REGION Network 7
   // *********************************************************************************************************************
   // 
   // Next Carrier Traffic Cop Motion Function Block FB111. Traffic Cop and carrier motion logic for Zone called in Function block call located  in OB1.  Function block contains logic for Motion control and Traffic Cop logic for Carrier located in Position 3 of called Zone.  Carrier position within the zone is contained in the Tag    - “ Zone.[called zone].CarrierZnStatus[Position in zone].  Input parameter “MaxCarriers” Zones are divided into positions based on “MaxCarriers” allowed in zone which is set in the zone setup function block and represents the maximum number of carriers within the zone. 
   // 
   // **********************************************************************************************************************
   RUNG wire#powerrail
      "IDB602_NextCarrierTCopMotionFB"(Zone := #Zone, ZonePos := 3, CarrierNumber => "DB116_TC_ZoneMotionControl".Zone[#Zone].ZonePos[3].CarrierNumber, MoveFwdCommand => "DB116_TC_ZoneMotionControl".Zone[#Zone].ZonePos[3].MoveFwd, DriveCmdSpeed => "DB116_TC_ZoneMotionControl".Zone[#Zone].ZonePos[3].DriveCmdSpeed, NextStopPosition => "DB116_TC_ZoneMotionControl".Zone[#Zone].ZonePos[3].NextStopPos, NextCarrierNum => "DB116_TC_ZoneMotionControl".Zone[#Zone].ZonePos[3].NextCarrierNumber, AtCmdPosition => "DB116_TC_ZoneMotionControl".Zone[#Zone].ZonePos[3].AtCmdPos)
   END_RUNG
   // the same network as SCL:
   "IDB602_NextCarrierTCopMotionFB"(Zone := #Zone,   // "FB111_NextCarrierTCopMotionFB"
                           ZonePos := 3,
                           CarrierNumber => "DB116_TC_ZoneMotionControl".Zone[#Zone].ZonePos[3].CarrierNumber,
                           MoveFwdCommand => "DB116_TC_ZoneMotionControl".Zone[#Zone].ZonePos[3].MoveFwd,
                           DriveCmdSpeed => "DB116_TC_ZoneMotionControl".Zone[#Zone].ZonePos[3].DriveCmdSpeed,
                           NextStopPosition => "DB116_TC_ZoneMotionControl".Zone[#Zone].ZonePos[3].NextStopPos,
                           NextCarrierNum => "DB116_TC_ZoneMotionControl".Zone[#Zone].ZonePos[3].NextCarrierNumber,
                           AtCmdPosition => "DB116_TC_ZoneMotionControl".Zone[#Zone].ZonePos[3].AtCmdPos);
END_REGION

REGION Network 8
   // *********************************************************************************************************************
   // 
   // Next Carrier Traffic Cop Motion Function Block FB111. Traffic Cop and carrier motion logic for Zone called in Function block call located  in OB1.  Function block contains logic for Motion control and Traffic Cop logic for Carrier located in Position 4 of called Zone.  Carrier position within the zone is contained in the Tag    - “ Zone.[called zone].CarrierZnStatus[Position in zone].  Input parameter “MaxCarriers” Zones are divided into positions based on “MaxCarriers” allowed in zone which is set in the zone setup function block and represents the maximum number of carriers within the zone. 
   // 
   // **********************************************************************************************************************
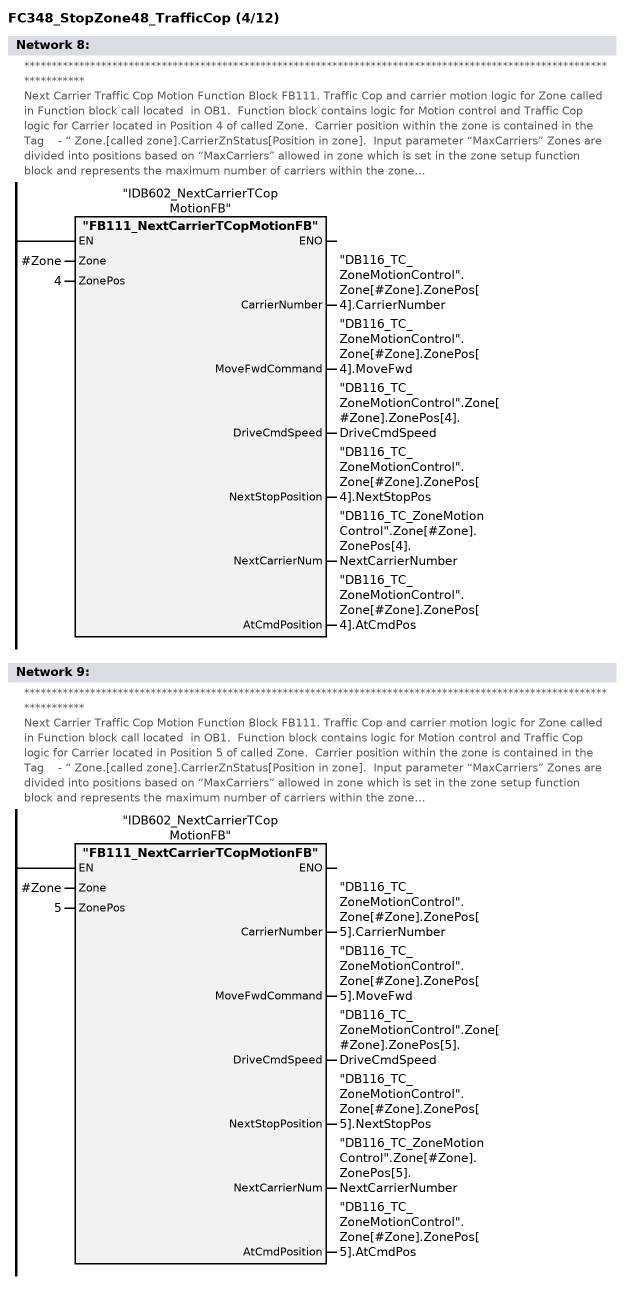
   RUNG wire#powerrail
      "IDB602_NextCarrierTCopMotionFB"(Zone := #Zone, ZonePos := 4, CarrierNumber => "DB116_TC_ZoneMotionControl".Zone[#Zone].ZonePos[4].CarrierNumber, MoveFwdCommand => "DB116_TC_ZoneMotionControl".Zone[#Zone].ZonePos[4].MoveFwd, DriveCmdSpeed => "DB116_TC_ZoneMotionControl".Zone[#Zone].ZonePos[4].DriveCmdSpeed, NextStopPosition => "DB116_TC_ZoneMotionControl".Zone[#Zone].ZonePos[4].NextStopPos, NextCarrierNum => "DB116_TC_ZoneMotionControl".Zone[#Zone].ZonePos[4].NextCarrierNumber, AtCmdPosition => "DB116_TC_ZoneMotionControl".Zone[#Zone].ZonePos[4].AtCmdPos)
   END_RUNG
   // the same network as SCL:
   "IDB602_NextCarrierTCopMotionFB"(Zone := #Zone,   // "FB111_NextCarrierTCopMotionFB"
                           ZonePos := 4,
                           CarrierNumber => "DB116_TC_ZoneMotionControl".Zone[#Zone].ZonePos[4].CarrierNumber,
                           MoveFwdCommand => "DB116_TC_ZoneMotionControl".Zone[#Zone].ZonePos[4].MoveFwd,
                           DriveCmdSpeed => "DB116_TC_ZoneMotionControl".Zone[#Zone].ZonePos[4].DriveCmdSpeed,
                           NextStopPosition => "DB116_TC_ZoneMotionControl".Zone[#Zone].ZonePos[4].NextStopPos,
                           NextCarrierNum => "DB116_TC_ZoneMotionControl".Zone[#Zone].ZonePos[4].NextCarrierNumber,
                           AtCmdPosition => "DB116_TC_ZoneMotionControl".Zone[#Zone].ZonePos[4].AtCmdPos);
END_REGION

REGION Network 9
   // *********************************************************************************************************************
   // 
   // Next Carrier Traffic Cop Motion Function Block FB111. Traffic Cop and carrier motion logic for Zone called in Function block call located  in OB1.  Function block contains logic for Motion control and Traffic Cop logic for Carrier located in Position 5 of called Zone.  Carrier position within the zone is contained in the Tag    - “ Zone.[called zone].CarrierZnStatus[Position in zone].  Input parameter “MaxCarriers” Zones are divided into positions based on “MaxCarriers” allowed in zone which is set in the zone setup function block and represents the maximum number of carriers within the zone. 
   // 
   // **********************************************************************************************************************
   RUNG wire#powerrail
      "IDB602_NextCarrierTCopMotionFB"(Zone := #Zone, ZonePos := 5, CarrierNumber => "DB116_TC_ZoneMotionControl".Zone[#Zone].ZonePos[5].CarrierNumber, MoveFwdCommand => "DB116_TC_ZoneMotionControl".Zone[#Zone].ZonePos[5].MoveFwd, DriveCmdSpeed => "DB116_TC_ZoneMotionControl".Zone[#Zone].ZonePos[5].DriveCmdSpeed, NextStopPosition => "DB116_TC_ZoneMotionControl".Zone[#Zone].ZonePos[5].NextStopPos, NextCarrierNum => "DB116_TC_ZoneMotionControl".Zone[#Zone].ZonePos[5].NextCarrierNumber, AtCmdPosition => "DB116_TC_ZoneMotionControl".Zone[#Zone].ZonePos[5].AtCmdPos)
   END_RUNG
   // the same network as SCL:
   "IDB602_NextCarrierTCopMotionFB"(Zone := #Zone,   // "FB111_NextCarrierTCopMotionFB"
                           ZonePos := 5,
                           CarrierNumber => "DB116_TC_ZoneMotionControl".Zone[#Zone].ZonePos[5].CarrierNumber,
                           MoveFwdCommand => "DB116_TC_ZoneMotionControl".Zone[#Zone].ZonePos[5].MoveFwd,
                           DriveCmdSpeed => "DB116_TC_ZoneMotionControl".Zone[#Zone].ZonePos[5].DriveCmdSpeed,
                           NextStopPosition => "DB116_TC_ZoneMotionControl".Zone[#Zone].ZonePos[5].NextStopPos,
                           NextCarrierNum => "DB116_TC_ZoneMotionControl".Zone[#Zone].ZonePos[5].NextCarrierNumber,
                           AtCmdPosition => "DB116_TC_ZoneMotionControl".Zone[#Zone].ZonePos[5].AtCmdPos);
END_REGION

REGION Network 10
   // *********************************************************************************************************************
   // 
   // Next Carrier Traffic Cop Motion Function Block FB111. Traffic Cop and carrier motion logic for Zone called in Function block call located  in OB1.  Function block contains logic for Motion control and Traffic Cop logic for Carrier located in Position 6 of called Zone.  Carrier position within the zone is contained in the Tag    - “ Zone.[called zone].CarrierZnStatus[Position in zone].  Input parameter “MaxCarriers” Zones are divided into positions based on “MaxCarriers” allowed in zone which is set in the zone setup function block and represents the maximum number of carriers within the zone. 
   // 
   // **********************************************************************************************************************
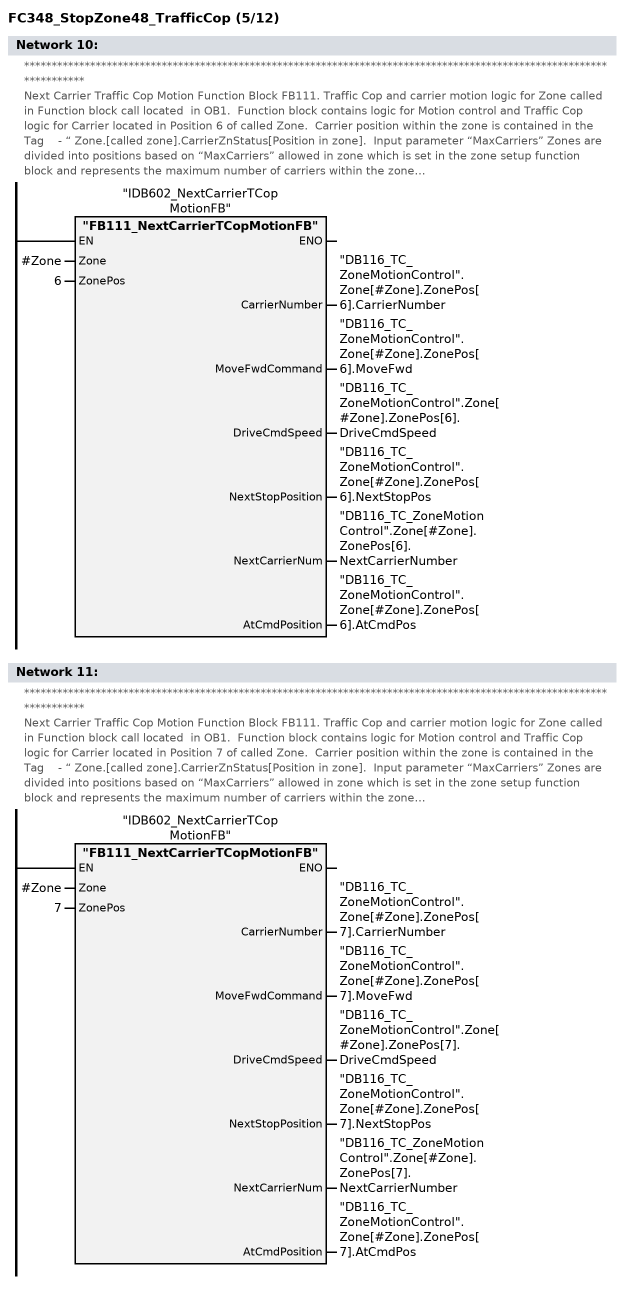
   RUNG wire#powerrail
      "IDB602_NextCarrierTCopMotionFB"(Zone := #Zone, ZonePos := 6, CarrierNumber => "DB116_TC_ZoneMotionControl".Zone[#Zone].ZonePos[6].CarrierNumber, MoveFwdCommand => "DB116_TC_ZoneMotionControl".Zone[#Zone].ZonePos[6].MoveFwd, DriveCmdSpeed => "DB116_TC_ZoneMotionControl".Zone[#Zone].ZonePos[6].DriveCmdSpeed, NextStopPosition => "DB116_TC_ZoneMotionControl".Zone[#Zone].ZonePos[6].NextStopPos, NextCarrierNum => "DB116_TC_ZoneMotionControl".Zone[#Zone].ZonePos[6].NextCarrierNumber, AtCmdPosition => "DB116_TC_ZoneMotionControl".Zone[#Zone].ZonePos[6].AtCmdPos)
   END_RUNG
   // the same network as SCL:
   "IDB602_NextCarrierTCopMotionFB"(Zone := #Zone,   // "FB111_NextCarrierTCopMotionFB"
                           ZonePos := 6,
                           CarrierNumber => "DB116_TC_ZoneMotionControl".Zone[#Zone].ZonePos[6].CarrierNumber,
                           MoveFwdCommand => "DB116_TC_ZoneMotionControl".Zone[#Zone].ZonePos[6].MoveFwd,
                           DriveCmdSpeed => "DB116_TC_ZoneMotionControl".Zone[#Zone].ZonePos[6].DriveCmdSpeed,
                           NextStopPosition => "DB116_TC_ZoneMotionControl".Zone[#Zone].ZonePos[6].NextStopPos,
                           NextCarrierNum => "DB116_TC_ZoneMotionControl".Zone[#Zone].ZonePos[6].NextCarrierNumber,
                           AtCmdPosition => "DB116_TC_ZoneMotionControl".Zone[#Zone].ZonePos[6].AtCmdPos);
END_REGION

REGION Network 11
   // *********************************************************************************************************************
   // 
   // Next Carrier Traffic Cop Motion Function Block FB111. Traffic Cop and carrier motion logic for Zone called in Function block call located  in OB1.  Function block contains logic for Motion control and Traffic Cop logic for Carrier located in Position 7 of called Zone.  Carrier position within the zone is contained in the Tag    - “ Zone.[called zone].CarrierZnStatus[Position in zone].  Input parameter “MaxCarriers” Zones are divided into positions based on “MaxCarriers” allowed in zone which is set in the zone setup function block and represents the maximum number of carriers within the zone. 
   // 
   // **********************************************************************************************************************
   RUNG wire#powerrail
      "IDB602_NextCarrierTCopMotionFB"(Zone := #Zone, ZonePos := 7, CarrierNumber => "DB116_TC_ZoneMotionControl".Zone[#Zone].ZonePos[7].CarrierNumber, MoveFwdCommand => "DB116_TC_ZoneMotionControl".Zone[#Zone].ZonePos[7].MoveFwd, DriveCmdSpeed => "DB116_TC_ZoneMotionControl".Zone[#Zone].ZonePos[7].DriveCmdSpeed, NextStopPosition => "DB116_TC_ZoneMotionControl".Zone[#Zone].ZonePos[7].NextStopPos, NextCarrierNum => "DB116_TC_ZoneMotionControl".Zone[#Zone].ZonePos[7].NextCarrierNumber, AtCmdPosition => "DB116_TC_ZoneMotionControl".Zone[#Zone].ZonePos[7].AtCmdPos)
   END_RUNG
   // the same network as SCL:
   "IDB602_NextCarrierTCopMotionFB"(Zone := #Zone,   // "FB111_NextCarrierTCopMotionFB"
                           ZonePos := 7,
                           CarrierNumber => "DB116_TC_ZoneMotionControl".Zone[#Zone].ZonePos[7].CarrierNumber,
                           MoveFwdCommand => "DB116_TC_ZoneMotionControl".Zone[#Zone].ZonePos[7].MoveFwd,
                           DriveCmdSpeed => "DB116_TC_ZoneMotionControl".Zone[#Zone].ZonePos[7].DriveCmdSpeed,
                           NextStopPosition => "DB116_TC_ZoneMotionControl".Zone[#Zone].ZonePos[7].NextStopPos,
                           NextCarrierNum => "DB116_TC_ZoneMotionControl".Zone[#Zone].ZonePos[7].NextCarrierNumber,
                           AtCmdPosition => "DB116_TC_ZoneMotionControl".Zone[#Zone].ZonePos[7].AtCmdPos);
END_REGION

REGION Network 12
   // *********************************************************************************************************************
   // 
   // Next Carrier Traffic Cop Motion Function Block FB111. Traffic Cop and carrier motion logic for Zone called in Function block call located  in OB1.  Function block contains logic for Motion control and Traffic Cop logic for Carrier located in Position 8 of called Zone.  Carrier position within the zone is contained in the Tag    - “ Zone.[called zone].CarrierZnStatus[Position in zone].  Input parameter “MaxCarriers” Zones are divided into positions based on “MaxCarriers” allowed in zone which is set in the zone setup function block and represents the maximum number of carriers within the zone. 
   // 
   // **********************************************************************************************************************
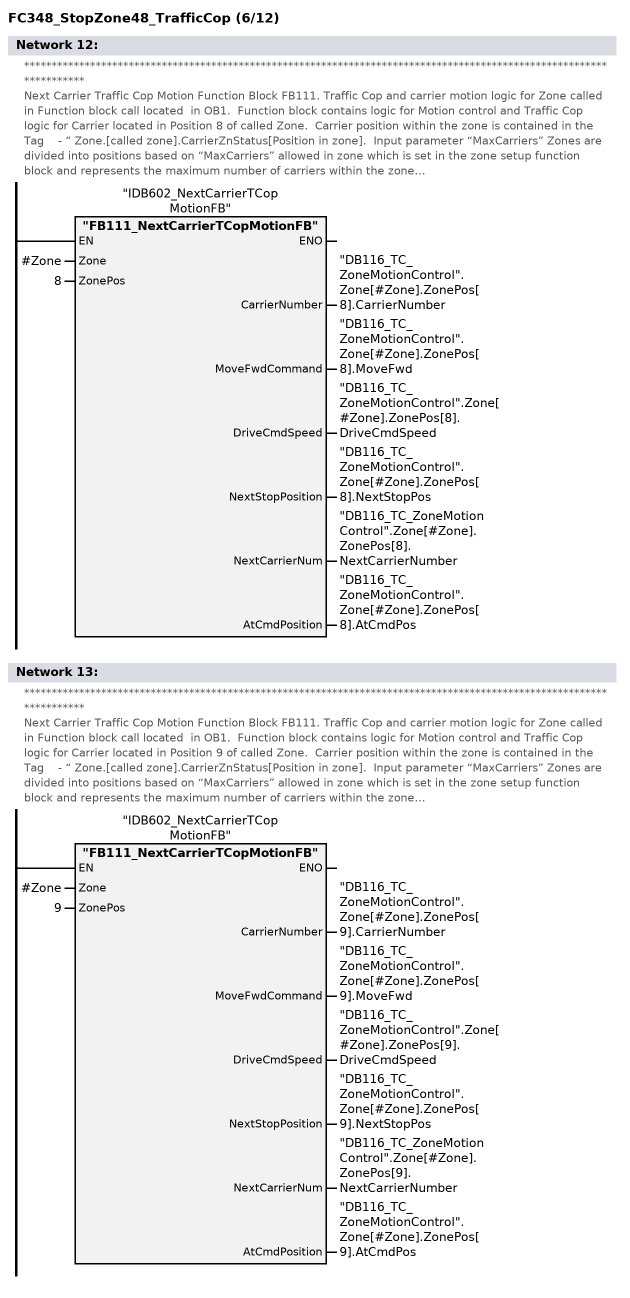
   RUNG wire#powerrail
      "IDB602_NextCarrierTCopMotionFB"(Zone := #Zone, ZonePos := 8, CarrierNumber => "DB116_TC_ZoneMotionControl".Zone[#Zone].ZonePos[8].CarrierNumber, MoveFwdCommand => "DB116_TC_ZoneMotionControl".Zone[#Zone].ZonePos[8].MoveFwd, DriveCmdSpeed => "DB116_TC_ZoneMotionControl".Zone[#Zone].ZonePos[8].DriveCmdSpeed, NextStopPosition => "DB116_TC_ZoneMotionControl".Zone[#Zone].ZonePos[8].NextStopPos, NextCarrierNum => "DB116_TC_ZoneMotionControl".Zone[#Zone].ZonePos[8].NextCarrierNumber, AtCmdPosition => "DB116_TC_ZoneMotionControl".Zone[#Zone].ZonePos[8].AtCmdPos)
   END_RUNG
   // the same network as SCL:
   "IDB602_NextCarrierTCopMotionFB"(Zone := #Zone,   // "FB111_NextCarrierTCopMotionFB"
                           ZonePos := 8,
                           CarrierNumber => "DB116_TC_ZoneMotionControl".Zone[#Zone].ZonePos[8].CarrierNumber,
                           MoveFwdCommand => "DB116_TC_ZoneMotionControl".Zone[#Zone].ZonePos[8].MoveFwd,
                           DriveCmdSpeed => "DB116_TC_ZoneMotionControl".Zone[#Zone].ZonePos[8].DriveCmdSpeed,
                           NextStopPosition => "DB116_TC_ZoneMotionControl".Zone[#Zone].ZonePos[8].NextStopPos,
                           NextCarrierNum => "DB116_TC_ZoneMotionControl".Zone[#Zone].ZonePos[8].NextCarrierNumber,
                           AtCmdPosition => "DB116_TC_ZoneMotionControl".Zone[#Zone].ZonePos[8].AtCmdPos);
END_REGION

REGION Network 13
   // *********************************************************************************************************************
   // 
   // Next Carrier Traffic Cop Motion Function Block FB111. Traffic Cop and carrier motion logic for Zone called in Function block call located  in OB1.  Function block contains logic for Motion control and Traffic Cop logic for Carrier located in Position 9 of called Zone.  Carrier position within the zone is contained in the Tag    - “ Zone.[called zone].CarrierZnStatus[Position in zone].  Input parameter “MaxCarriers” Zones are divided into positions based on “MaxCarriers” allowed in zone which is set in the zone setup function block and represents the maximum number of carriers within the zone. 
   // 
   // **********************************************************************************************************************
   RUNG wire#powerrail
      "IDB602_NextCarrierTCopMotionFB"(Zone := #Zone, ZonePos := 9, CarrierNumber => "DB116_TC_ZoneMotionControl".Zone[#Zone].ZonePos[9].CarrierNumber, MoveFwdCommand => "DB116_TC_ZoneMotionControl".Zone[#Zone].ZonePos[9].MoveFwd, DriveCmdSpeed => "DB116_TC_ZoneMotionControl".Zone[#Zone].ZonePos[9].DriveCmdSpeed, NextStopPosition => "DB116_TC_ZoneMotionControl".Zone[#Zone].ZonePos[9].NextStopPos, NextCarrierNum => "DB116_TC_ZoneMotionControl".Zone[#Zone].ZonePos[9].NextCarrierNumber, AtCmdPosition => "DB116_TC_ZoneMotionControl".Zone[#Zone].ZonePos[9].AtCmdPos)
   END_RUNG
   // the same network as SCL:
   "IDB602_NextCarrierTCopMotionFB"(Zone := #Zone,   // "FB111_NextCarrierTCopMotionFB"
                           ZonePos := 9,
                           CarrierNumber => "DB116_TC_ZoneMotionControl".Zone[#Zone].ZonePos[9].CarrierNumber,
                           MoveFwdCommand => "DB116_TC_ZoneMotionControl".Zone[#Zone].ZonePos[9].MoveFwd,
                           DriveCmdSpeed => "DB116_TC_ZoneMotionControl".Zone[#Zone].ZonePos[9].DriveCmdSpeed,
                           NextStopPosition => "DB116_TC_ZoneMotionControl".Zone[#Zone].ZonePos[9].NextStopPos,
                           NextCarrierNum => "DB116_TC_ZoneMotionControl".Zone[#Zone].ZonePos[9].NextCarrierNumber,
                           AtCmdPosition => "DB116_TC_ZoneMotionControl".Zone[#Zone].ZonePos[9].AtCmdPos);
END_REGION

REGION Network 14
   // *********************************************************************************************************************
   // 
   // Next Carrier Traffic Cop Motion Function Block FB111. Traffic Cop and carrier motion logic for Zone called in Function block call located  in OB1.  Function block contains logic for Motion control and Traffic Cop logic for Carrier located in Position 10 of called Zone.  Carrier position within the zone is contained in the Tag    - “ Zone.[called zone].CarrierZnStatus[Position in zone].  Input parameter “MaxCarriers” Zones are divided into positions based on “MaxCarriers” allowed in zone which is set in the zone setup function block and represents the maximum number of carriers within the zone. 
   // 
   // **********************************************************************************************************************
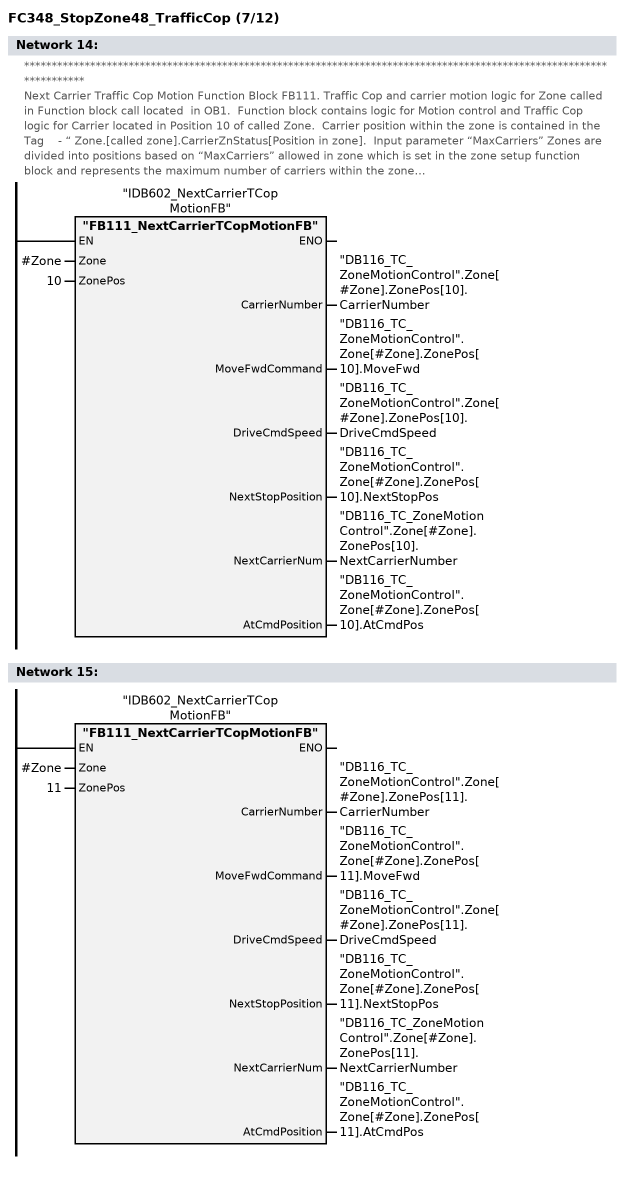
   RUNG wire#powerrail
      "IDB602_NextCarrierTCopMotionFB"(Zone := #Zone, ZonePos := 10, CarrierNumber => "DB116_TC_ZoneMotionControl".Zone[#Zone].ZonePos[10].CarrierNumber, MoveFwdCommand => "DB116_TC_ZoneMotionControl".Zone[#Zone].ZonePos[10].MoveFwd, DriveCmdSpeed => "DB116_TC_ZoneMotionControl".Zone[#Zone].ZonePos[10].DriveCmdSpeed, NextStopPosition => "DB116_TC_ZoneMotionControl".Zone[#Zone].ZonePos[10].NextStopPos, NextCarrierNum => "DB116_TC_ZoneMotionControl".Zone[#Zone].ZonePos[10].NextCarrierNumber, AtCmdPosition => "DB116_TC_ZoneMotionControl".Zone[#Zone].ZonePos[10].AtCmdPos)
   END_RUNG
   // the same network as SCL:
   "IDB602_NextCarrierTCopMotionFB"(Zone := #Zone,   // "FB111_NextCarrierTCopMotionFB"
                           ZonePos := 10,
                           CarrierNumber => "DB116_TC_ZoneMotionControl".Zone[#Zone].ZonePos[10].CarrierNumber,
                           MoveFwdCommand => "DB116_TC_ZoneMotionControl".Zone[#Zone].ZonePos[10].MoveFwd,
                           DriveCmdSpeed => "DB116_TC_ZoneMotionControl".Zone[#Zone].ZonePos[10].DriveCmdSpeed,
                           NextStopPosition => "DB116_TC_ZoneMotionControl".Zone[#Zone].ZonePos[10].NextStopPos,
                           NextCarrierNum => "DB116_TC_ZoneMotionControl".Zone[#Zone].ZonePos[10].NextCarrierNumber,
                           AtCmdPosition => "DB116_TC_ZoneMotionControl".Zone[#Zone].ZonePos[10].AtCmdPos);
END_REGION

REGION Network 15
   RUNG wire#powerrail
      "IDB602_NextCarrierTCopMotionFB"(Zone := #Zone, ZonePos := 11, CarrierNumber => "DB116_TC_ZoneMotionControl".Zone[#Zone].ZonePos[11].CarrierNumber, MoveFwdCommand => "DB116_TC_ZoneMotionControl".Zone[#Zone].ZonePos[11].MoveFwd, DriveCmdSpeed => "DB116_TC_ZoneMotionControl".Zone[#Zone].ZonePos[11].DriveCmdSpeed, NextStopPosition => "DB116_TC_ZoneMotionControl".Zone[#Zone].ZonePos[11].NextStopPos, NextCarrierNum => "DB116_TC_ZoneMotionControl".Zone[#Zone].ZonePos[11].NextCarrierNumber, AtCmdPosition => "DB116_TC_ZoneMotionControl".Zone[#Zone].ZonePos[11].AtCmdPos)
   END_RUNG
   // the same network as SCL:
   "IDB602_NextCarrierTCopMotionFB"(Zone := #Zone,   // "FB111_NextCarrierTCopMotionFB"
                           ZonePos := 11,
                           CarrierNumber => "DB116_TC_ZoneMotionControl".Zone[#Zone].ZonePos[11].CarrierNumber,
                           MoveFwdCommand => "DB116_TC_ZoneMotionControl".Zone[#Zone].ZonePos[11].MoveFwd,
                           DriveCmdSpeed => "DB116_TC_ZoneMotionControl".Zone[#Zone].ZonePos[11].DriveCmdSpeed,
                           NextStopPosition => "DB116_TC_ZoneMotionControl".Zone[#Zone].ZonePos[11].NextStopPos,
                           NextCarrierNum => "DB116_TC_ZoneMotionControl".Zone[#Zone].ZonePos[11].NextCarrierNumber,
                           AtCmdPosition => "DB116_TC_ZoneMotionControl".Zone[#Zone].ZonePos[11].AtCmdPos);
END_REGION

REGION Network 16
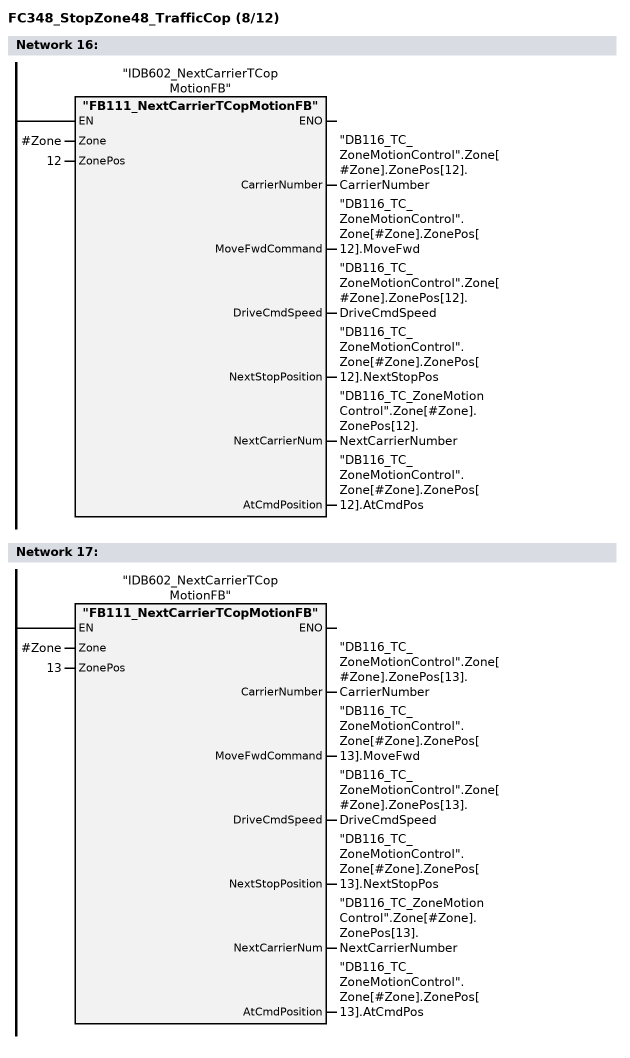
   RUNG wire#powerrail
      "IDB602_NextCarrierTCopMotionFB"(Zone := #Zone, ZonePos := 12, CarrierNumber => "DB116_TC_ZoneMotionControl".Zone[#Zone].ZonePos[12].CarrierNumber, MoveFwdCommand => "DB116_TC_ZoneMotionControl".Zone[#Zone].ZonePos[12].MoveFwd, DriveCmdSpeed => "DB116_TC_ZoneMotionControl".Zone[#Zone].ZonePos[12].DriveCmdSpeed, NextStopPosition => "DB116_TC_ZoneMotionControl".Zone[#Zone].ZonePos[12].NextStopPos, NextCarrierNum => "DB116_TC_ZoneMotionControl".Zone[#Zone].ZonePos[12].NextCarrierNumber, AtCmdPosition => "DB116_TC_ZoneMotionControl".Zone[#Zone].ZonePos[12].AtCmdPos)
   END_RUNG
   // the same network as SCL:
   "IDB602_NextCarrierTCopMotionFB"(Zone := #Zone,   // "FB111_NextCarrierTCopMotionFB"
                           ZonePos := 12,
                           CarrierNumber => "DB116_TC_ZoneMotionControl".Zone[#Zone].ZonePos[12].CarrierNumber,
                           MoveFwdCommand => "DB116_TC_ZoneMotionControl".Zone[#Zone].ZonePos[12].MoveFwd,
                           DriveCmdSpeed => "DB116_TC_ZoneMotionControl".Zone[#Zone].ZonePos[12].DriveCmdSpeed,
                           NextStopPosition => "DB116_TC_ZoneMotionControl".Zone[#Zone].ZonePos[12].NextStopPos,
                           NextCarrierNum => "DB116_TC_ZoneMotionControl".Zone[#Zone].ZonePos[12].NextCarrierNumber,
                           AtCmdPosition => "DB116_TC_ZoneMotionControl".Zone[#Zone].ZonePos[12].AtCmdPos);
END_REGION

REGION Network 17
   RUNG wire#powerrail
      "IDB602_NextCarrierTCopMotionFB"(Zone := #Zone, ZonePos := 13, CarrierNumber => "DB116_TC_ZoneMotionControl".Zone[#Zone].ZonePos[13].CarrierNumber, MoveFwdCommand => "DB116_TC_ZoneMotionControl".Zone[#Zone].ZonePos[13].MoveFwd, DriveCmdSpeed => "DB116_TC_ZoneMotionControl".Zone[#Zone].ZonePos[13].DriveCmdSpeed, NextStopPosition => "DB116_TC_ZoneMotionControl".Zone[#Zone].ZonePos[13].NextStopPos, NextCarrierNum => "DB116_TC_ZoneMotionControl".Zone[#Zone].ZonePos[13].NextCarrierNumber, AtCmdPosition => "DB116_TC_ZoneMotionControl".Zone[#Zone].ZonePos[13].AtCmdPos)
   END_RUNG
   // the same network as SCL:
   "IDB602_NextCarrierTCopMotionFB"(Zone := #Zone,   // "FB111_NextCarrierTCopMotionFB"
                           ZonePos := 13,
                           CarrierNumber => "DB116_TC_ZoneMotionControl".Zone[#Zone].ZonePos[13].CarrierNumber,
                           MoveFwdCommand => "DB116_TC_ZoneMotionControl".Zone[#Zone].ZonePos[13].MoveFwd,
                           DriveCmdSpeed => "DB116_TC_ZoneMotionControl".Zone[#Zone].ZonePos[13].DriveCmdSpeed,
                           NextStopPosition => "DB116_TC_ZoneMotionControl".Zone[#Zone].ZonePos[13].NextStopPos,
                           NextCarrierNum => "DB116_TC_ZoneMotionControl".Zone[#Zone].ZonePos[13].NextCarrierNumber,
                           AtCmdPosition => "DB116_TC_ZoneMotionControl".Zone[#Zone].ZonePos[13].AtCmdPos);
END_REGION

REGION Network 18
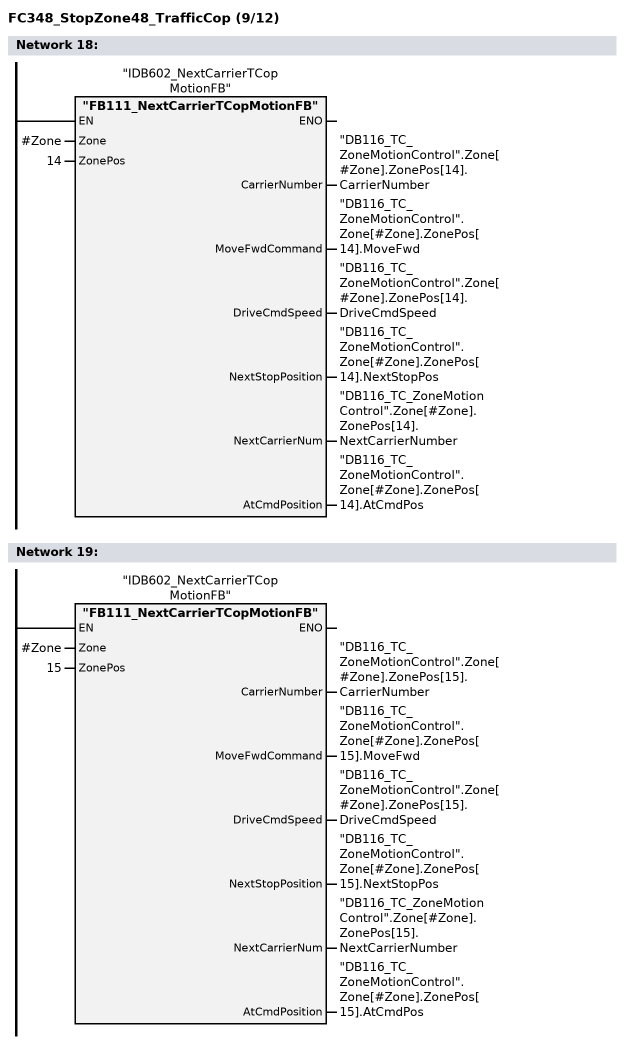
   RUNG wire#powerrail
      "IDB602_NextCarrierTCopMotionFB"(Zone := #Zone, ZonePos := 14, CarrierNumber => "DB116_TC_ZoneMotionControl".Zone[#Zone].ZonePos[14].CarrierNumber, MoveFwdCommand => "DB116_TC_ZoneMotionControl".Zone[#Zone].ZonePos[14].MoveFwd, DriveCmdSpeed => "DB116_TC_ZoneMotionControl".Zone[#Zone].ZonePos[14].DriveCmdSpeed, NextStopPosition => "DB116_TC_ZoneMotionControl".Zone[#Zone].ZonePos[14].NextStopPos, NextCarrierNum => "DB116_TC_ZoneMotionControl".Zone[#Zone].ZonePos[14].NextCarrierNumber, AtCmdPosition => "DB116_TC_ZoneMotionControl".Zone[#Zone].ZonePos[14].AtCmdPos)
   END_RUNG
   // the same network as SCL:
   "IDB602_NextCarrierTCopMotionFB"(Zone := #Zone,   // "FB111_NextCarrierTCopMotionFB"
                           ZonePos := 14,
                           CarrierNumber => "DB116_TC_ZoneMotionControl".Zone[#Zone].ZonePos[14].CarrierNumber,
                           MoveFwdCommand => "DB116_TC_ZoneMotionControl".Zone[#Zone].ZonePos[14].MoveFwd,
                           DriveCmdSpeed => "DB116_TC_ZoneMotionControl".Zone[#Zone].ZonePos[14].DriveCmdSpeed,
                           NextStopPosition => "DB116_TC_ZoneMotionControl".Zone[#Zone].ZonePos[14].NextStopPos,
                           NextCarrierNum => "DB116_TC_ZoneMotionControl".Zone[#Zone].ZonePos[14].NextCarrierNumber,
                           AtCmdPosition => "DB116_TC_ZoneMotionControl".Zone[#Zone].ZonePos[14].AtCmdPos);
END_REGION

REGION Network 19
   RUNG wire#powerrail
      "IDB602_NextCarrierTCopMotionFB"(Zone := #Zone, ZonePos := 15, CarrierNumber => "DB116_TC_ZoneMotionControl".Zone[#Zone].ZonePos[15].CarrierNumber, MoveFwdCommand => "DB116_TC_ZoneMotionControl".Zone[#Zone].ZonePos[15].MoveFwd, DriveCmdSpeed => "DB116_TC_ZoneMotionControl".Zone[#Zone].ZonePos[15].DriveCmdSpeed, NextStopPosition => "DB116_TC_ZoneMotionControl".Zone[#Zone].ZonePos[15].NextStopPos, NextCarrierNum => "DB116_TC_ZoneMotionControl".Zone[#Zone].ZonePos[15].NextCarrierNumber, AtCmdPosition => "DB116_TC_ZoneMotionControl".Zone[#Zone].ZonePos[15].AtCmdPos)
   END_RUNG
   // the same network as SCL:
   "IDB602_NextCarrierTCopMotionFB"(Zone := #Zone,   // "FB111_NextCarrierTCopMotionFB"
                           ZonePos := 15,
                           CarrierNumber => "DB116_TC_ZoneMotionControl".Zone[#Zone].ZonePos[15].CarrierNumber,
                           MoveFwdCommand => "DB116_TC_ZoneMotionControl".Zone[#Zone].ZonePos[15].MoveFwd,
                           DriveCmdSpeed => "DB116_TC_ZoneMotionControl".Zone[#Zone].ZonePos[15].DriveCmdSpeed,
                           NextStopPosition => "DB116_TC_ZoneMotionControl".Zone[#Zone].ZonePos[15].NextStopPos,
                           NextCarrierNum => "DB116_TC_ZoneMotionControl".Zone[#Zone].ZonePos[15].NextCarrierNumber,
                           AtCmdPosition => "DB116_TC_ZoneMotionControl".Zone[#Zone].ZonePos[15].AtCmdPos);
END_REGION

REGION Network 20
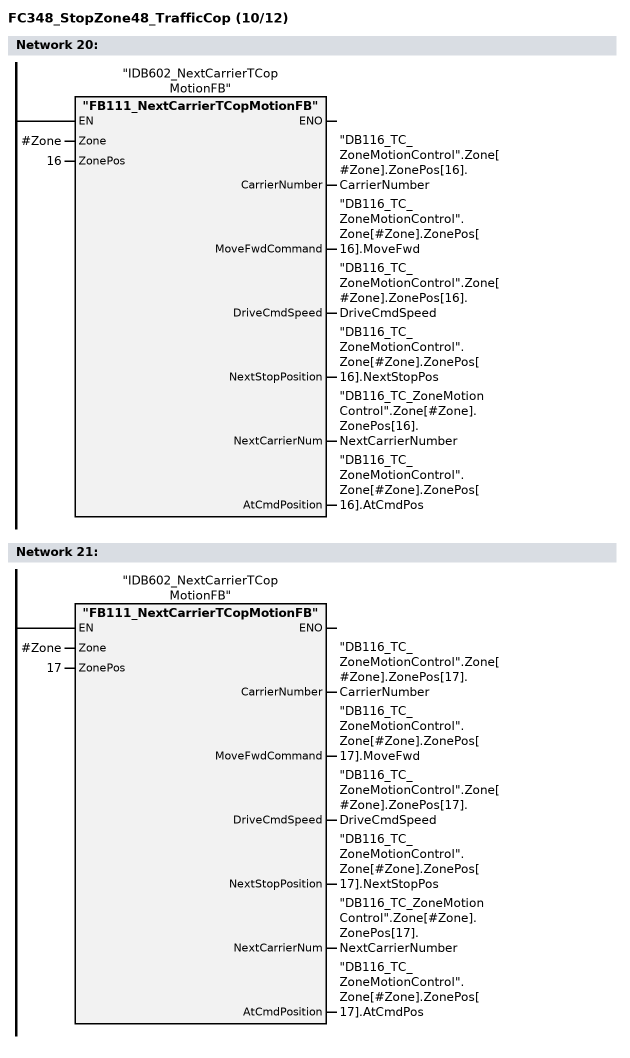
   RUNG wire#powerrail
      "IDB602_NextCarrierTCopMotionFB"(Zone := #Zone, ZonePos := 16, CarrierNumber => "DB116_TC_ZoneMotionControl".Zone[#Zone].ZonePos[16].CarrierNumber, MoveFwdCommand => "DB116_TC_ZoneMotionControl".Zone[#Zone].ZonePos[16].MoveFwd, DriveCmdSpeed => "DB116_TC_ZoneMotionControl".Zone[#Zone].ZonePos[16].DriveCmdSpeed, NextStopPosition => "DB116_TC_ZoneMotionControl".Zone[#Zone].ZonePos[16].NextStopPos, NextCarrierNum => "DB116_TC_ZoneMotionControl".Zone[#Zone].ZonePos[16].NextCarrierNumber, AtCmdPosition => "DB116_TC_ZoneMotionControl".Zone[#Zone].ZonePos[16].AtCmdPos)
   END_RUNG
   // the same network as SCL:
   "IDB602_NextCarrierTCopMotionFB"(Zone := #Zone,   // "FB111_NextCarrierTCopMotionFB"
                           ZonePos := 16,
                           CarrierNumber => "DB116_TC_ZoneMotionControl".Zone[#Zone].ZonePos[16].CarrierNumber,
                           MoveFwdCommand => "DB116_TC_ZoneMotionControl".Zone[#Zone].ZonePos[16].MoveFwd,
                           DriveCmdSpeed => "DB116_TC_ZoneMotionControl".Zone[#Zone].ZonePos[16].DriveCmdSpeed,
                           NextStopPosition => "DB116_TC_ZoneMotionControl".Zone[#Zone].ZonePos[16].NextStopPos,
                           NextCarrierNum => "DB116_TC_ZoneMotionControl".Zone[#Zone].ZonePos[16].NextCarrierNumber,
                           AtCmdPosition => "DB116_TC_ZoneMotionControl".Zone[#Zone].ZonePos[16].AtCmdPos);
END_REGION

REGION Network 21
   RUNG wire#powerrail
      "IDB602_NextCarrierTCopMotionFB"(Zone := #Zone, ZonePos := 17, CarrierNumber => "DB116_TC_ZoneMotionControl".Zone[#Zone].ZonePos[17].CarrierNumber, MoveFwdCommand => "DB116_TC_ZoneMotionControl".Zone[#Zone].ZonePos[17].MoveFwd, DriveCmdSpeed => "DB116_TC_ZoneMotionControl".Zone[#Zone].ZonePos[17].DriveCmdSpeed, NextStopPosition => "DB116_TC_ZoneMotionControl".Zone[#Zone].ZonePos[17].NextStopPos, NextCarrierNum => "DB116_TC_ZoneMotionControl".Zone[#Zone].ZonePos[17].NextCarrierNumber, AtCmdPosition => "DB116_TC_ZoneMotionControl".Zone[#Zone].ZonePos[17].AtCmdPos)
   END_RUNG
   // the same network as SCL:
   "IDB602_NextCarrierTCopMotionFB"(Zone := #Zone,   // "FB111_NextCarrierTCopMotionFB"
                           ZonePos := 17,
                           CarrierNumber => "DB116_TC_ZoneMotionControl".Zone[#Zone].ZonePos[17].CarrierNumber,
                           MoveFwdCommand => "DB116_TC_ZoneMotionControl".Zone[#Zone].ZonePos[17].MoveFwd,
                           DriveCmdSpeed => "DB116_TC_ZoneMotionControl".Zone[#Zone].ZonePos[17].DriveCmdSpeed,
                           NextStopPosition => "DB116_TC_ZoneMotionControl".Zone[#Zone].ZonePos[17].NextStopPos,
                           NextCarrierNum => "DB116_TC_ZoneMotionControl".Zone[#Zone].ZonePos[17].NextCarrierNumber,
                           AtCmdPosition => "DB116_TC_ZoneMotionControl".Zone[#Zone].ZonePos[17].AtCmdPos);
END_REGION

REGION Network 22